(* Logix 5000 project; controller FV vendor 1 type 14 code 217 rev 31.11; software revision 31.00; part 8 of 63 *)
(* tags used below, declared in another part *)
   CWD : CHECKWORD_FLAGS;
   FR_B240 : INT[255];   // DEBOUNCE Debounce Flags
   FR_Delphi_I : DINT[60];
   FR_FILT_PR_PX : PlantItem;   // FILT_PR_PX
   FR_FILT_PR_PX_RawInput : ALIAS FOR RIO_Rack_2:3:I.Data.25;   // FR_FILT_PR_PX
   FR_FILT_TNK_PX : PlantItem;   // FILT_TNK_PX
   FR_FILT_TNK_PX_RawInput : ALIAS FOR RIO_Rack_2:3:I.Data.26;   // FR_FILT_TNK_PX
   FR_FILT_TNLN_PX : PlantItem;   // FILT_TNLN_PX
   FR_FILT_TNLN_PX_RawInput : ALIAS FOR RIO_Rack_2:3:I.Data.27;   // FR_FILT_TNLN_PX
   FR_FRV1_LP01 : PlantItem;   // FRV1_LP01
   FR_FRV1_LP01_RawInput : ALIAS FOR RIO_Rack_2:3:I.Data.13;   // FR_FRV1_LP01
   FR_FV26_HLP01 : PlantItem;   // FV26_HLP01
   FR_FV26_HLP01_RawInput : ALIAS FOR RIO_Rack_2:3:I.Data.0;   // FR_FV26_HLP01
   FR_FV26_LLP01 : PlantItem;   // FV26_LLP01
   FR_FV26_LLP01_RawInput : ALIAS FOR RIO_Rack_2:3:I.Data.1;   // FR_FV26_LLP01
   FR_FV27_HLP01 : PlantItem;   // FV27_HLP01
   FR_FV27_HLP01_RawInput : ALIAS FOR RIO_Rack_2:3:I.Data.2;   // FR_FV27_HLP01
   FR_FV27_LLP01 : PlantItem;   // FV27_LLP01
   FR_FV27_LLP01_RawInput : ALIAS FOR RIO_Rack_2:3:I.Data.3;   // FR_FV27_LLP01
   FR_FV28_HLP01 : PlantItem;   // FV28_HLP01
   FR_FV28_HLP01_RawInput : ALIAS FOR RIO_Rack_2:3:I.Data.4;   // FR_FV28_HLP01
   FR_FV28_LLP01 : PlantItem;   // FV28_LLP01
   FR_FV28_LLP01_RawInput : ALIAS FOR RIO_Rack_2:3:I.Data.5;   // FR_FV28_LLP01
   FR_FV29_HLP01 : PlantItem;   // FV29_HLP01
   FR_FV29_HLP01_RawInput : ALIAS FOR RIO_Rack_2:3:I.Data.6;   // FR_FV29_HLP01
   FR_FV29_LLP01 : PlantItem;   // FV29_LLP01
   FR_FV29_LLP01_RawInput : ALIAS FOR RIO_Rack_2:3:I.Data.7;   // FR_FV29_LLP01
   FR_FV30_HLP01 : PlantItem;   // FV30_HLP01
   FR_FV30_HLP01_RawInput : ALIAS FOR RIO_Rack_2:3:I.Data.8;   // FR_FV30_HLP01
   FR_FV30_LLP01 : PlantItem;   // FV30_LLP01
   FR_FV30_LLP01_RawInput : ALIAS FOR RIO_Rack_2:3:I.Data.9;   // FR_FV30_LLP01
   FR_FV31_HLP01 : PlantItem;   // FV31_HLP01
   FR_FV31_HLP01_RawInput : ALIAS FOR RIO_Rack_2:3:I.Data.10;   // FR_FV31_HLP01
   FR_FV31_LLP01 : PlantItem;   // FV31_LLP01
   FR_FV31_LLP01_RawInput : ALIAS FOR RIO_Rack_2:3:I.Data.11;   // FR_FV31_LLP01
   FR_R3_SW3_3 : PlantItem;   // R3_SW3_3
   FR_R3_SW3_3_RawInput : ALIAS FOR RIO_Rack_2:3:I.Data.14;   // FR_R3_SW3_3 FR_N14[109].2
   FR_T242 : TIMER[255];   // DEBOUNCE
   FR_T243 : TIMER[255];   // DEBOUNCE
   FR_VB4_LP01 : PlantItem;   // VB4_LP01
   FR_VB4_LP01_RawInput : ALIAS FOR RIO_Rack_2:3:I.Data.12;   // FR_VB4_LP01
   FR_YP1_CIPRET : PlantItem;   // YP1_CIPRET
   FR_YP1_CIPRET_RawInput : ALIAS FOR RIO_Rack_2:3:I.Data.24;   // FR_YP1_CIPRET
   FR_YP2_CIPRET : PlantItem;   // YP2_CIPRET
   FR_YP2_CIPRET_RawInput : ALIAS FOR RIO_Rack_2:3:I.Data.22;   // FR_YP2_CIPRET
   FR_YP3_CIPRET : PlantItem;   // YP3_CIPRET
   FR_YP3_CIPRET_RawInput : ALIAS FOR RIO_Rack_2:3:I.Data.23;   // FR_YP3_CIPRET
   One_Second_One_Scan : ALIAS FOR One_Second_1_scan;
(* FR_Common, continued *)

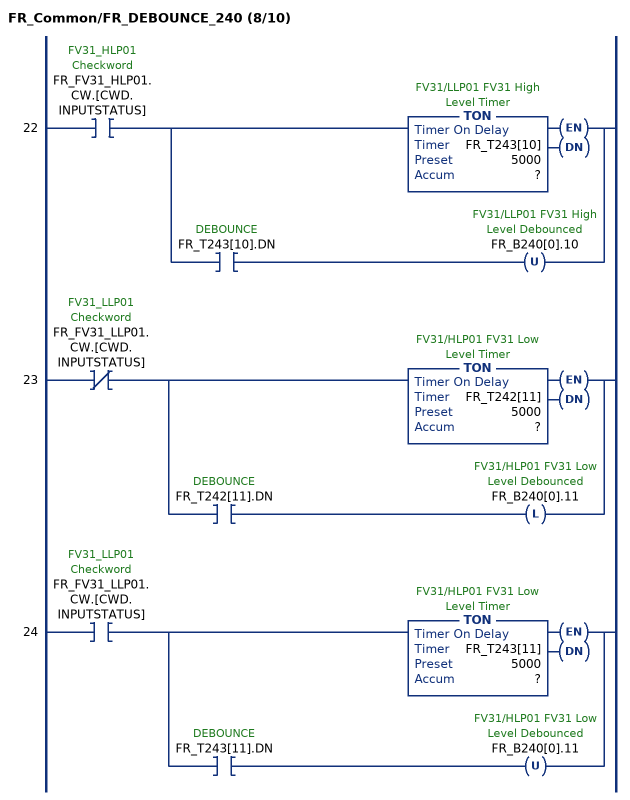
   [picture p70: FR_Common/FR_DEBOUNCE_240 rungs 22-24]
   22: XIC(FR_FV31_HLP01.CW.[CWD.INPUTSTATUS])[TON(FR_T243[10],?,?) ,XIC(FR_T243[10].DN) OTU(FR_B240[0].10) ];
   23: XIO(FR_FV31_LLP01.CW.[CWD.INPUTSTATUS])[TON(FR_T242[11],?,?) ,XIC(FR_T242[11].DN) OTL(FR_B240[0].11) ];
   24: XIC(FR_FV31_LLP01.CW.[CWD.INPUTSTATUS])[TON(FR_T243[11],?,?) ,XIC(FR_T243[11].DN) OTU(FR_B240[0].11) ];
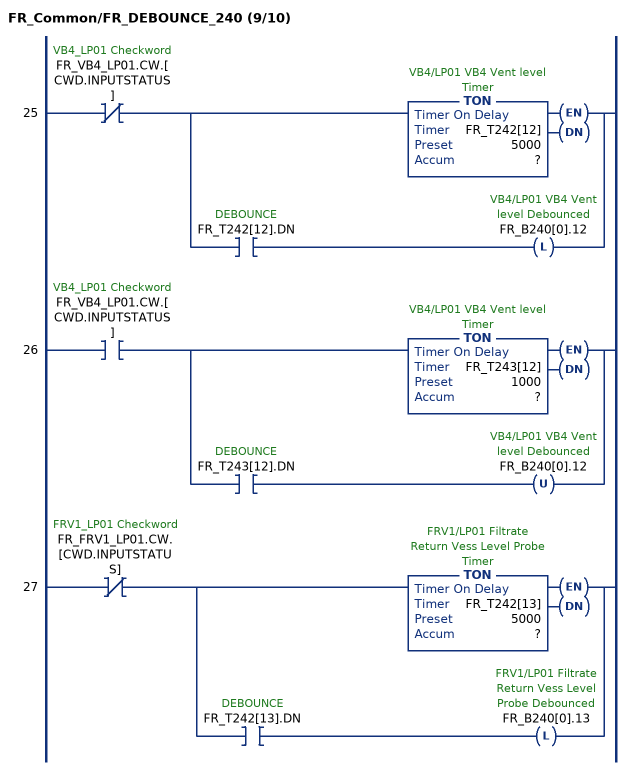
   25: XIO(FR_VB4_LP01.CW.[CWD.INPUTSTATUS])[TON(FR_T242[12],?,?) ,XIC(FR_T242[12].DN) OTL(FR_B240[0].12) ];
   26: XIC(FR_VB4_LP01.CW.[CWD.INPUTSTATUS])[TON(FR_T243[12],?,?) ,XIC(FR_T243[12].DN) OTU(FR_B240[0].12) ];
   27: XIO(FR_FRV1_LP01.CW.[CWD.INPUTSTATUS])[TON(FR_T242[13],?,?) ,XIC(FR_T242[13].DN) OTL(FR_B240[0].13) ];
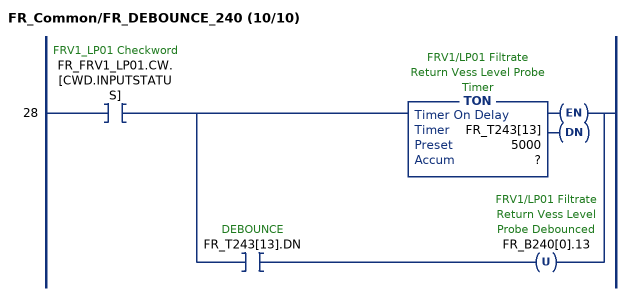
   28: XIC(FR_FRV1_LP01.CW.[CWD.INPUTSTATUS])[TON(FR_T243[13],?,?) ,XIC(FR_T243[13].DN) OTU(FR_B240[0].13) ];
END_ROUTINE

ROUTINE FR_Digital_Inputs   (* ladder *)
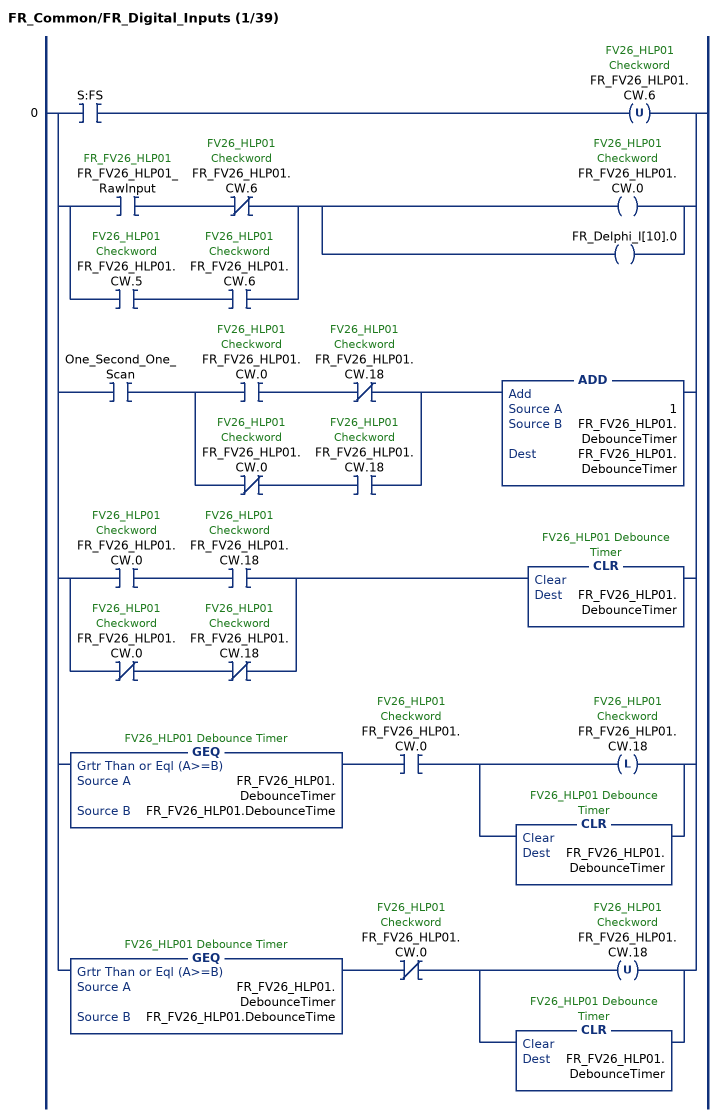
   0: [XIC(S:FS) OTU(FR_FV26_HLP01.CW.6) ,[XIC(FR_FV26_HLP01_RawInput) XIO(FR_FV26_HLP01.CW.6) ,XIC(FR_FV26_HLP01.CW.5) XIC(FR_FV26_HLP01.CW.6) ] [OTE(FR_FV26_HLP01.CW.0) ,OTE(FR_Delphi_I[10].0) ] ,XIC(One_Second_One_Scan) [XIC(FR_FV26_HLP01.CW.0) XIO(FR_FV26_HLP01.CW.18) ,XIO(FR_FV26_HLP01.CW.0) XIC(FR_FV26_HLP01.CW.18) ] ADD(1,FR_FV26_HLP01.DebounceTimer,FR_FV26_HLP01.DebounceTimer) ,[XIC(FR_FV26_HLP01.CW.0) XIC(FR_FV26_HLP01.CW.18) ,XIO(FR_FV26_HLP01.CW.0) XIO(FR_FV26_HLP01.CW.18) ] CLR(FR_FV26_HLP01.DebounceTimer) ,GEQ(FR_FV26_HLP01.DebounceTimer,FR_FV26_HLP01.DebounceTime) XIC(FR_FV26_HLP01.CW.0) [OTL(FR_FV26_HLP01.CW.18) ,CLR(FR_FV26_HLP01.DebounceTimer) ] ,GEQ(FR_FV26_HLP01.DebounceTimer,FR_FV26_HLP01.DebounceTime) XIO(FR_FV26_HLP01.CW.0) [OTU(FR_FV26_HLP01.CW.18) ,CLR(FR_FV26_HLP01.DebounceTimer) ] ];
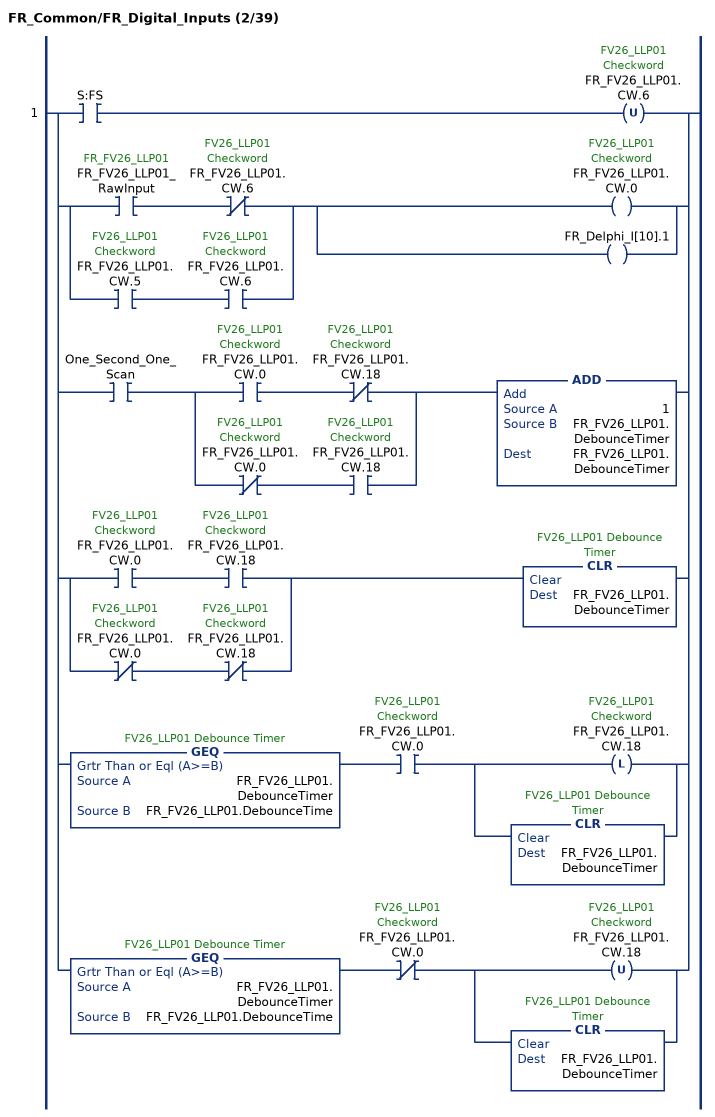
   1: [XIC(S:FS) OTU(FR_FV26_LLP01.CW.6) ,[XIC(FR_FV26_LLP01_RawInput) XIO(FR_FV26_LLP01.CW.6) ,XIC(FR_FV26_LLP01.CW.5) XIC(FR_FV26_LLP01.CW.6) ] [OTE(FR_FV26_LLP01.CW.0) ,OTE(FR_Delphi_I[10].1) ] ,XIC(One_Second_One_Scan) [XIC(FR_FV26_LLP01.CW.0) XIO(FR_FV26_LLP01.CW.18) ,XIO(FR_FV26_LLP01.CW.0) XIC(FR_FV26_LLP01.CW.18) ] ADD(1,FR_FV26_LLP01.DebounceTimer,FR_FV26_LLP01.DebounceTimer) ,[XIC(FR_FV26_LLP01.CW.0) XIC(FR_FV26_LLP01.CW.18) ,XIO(FR_FV26_LLP01.CW.0) XIO(FR_FV26_LLP01.CW.18) ] CLR(FR_FV26_LLP01.DebounceTimer) ,GEQ(FR_FV26_LLP01.DebounceTimer,FR_FV26_LLP01.DebounceTime) XIC(FR_FV26_LLP01.CW.0) [OTL(FR_FV26_LLP01.CW.18) ,CLR(FR_FV26_LLP01.DebounceTimer) ] ,GEQ(FR_FV26_LLP01.DebounceTimer,FR_FV26_LLP01.DebounceTime) XIO(FR_FV26_LLP01.CW.0) [OTU(FR_FV26_LLP01.CW.18) ,CLR(FR_FV26_LLP01.DebounceTimer) ] ];
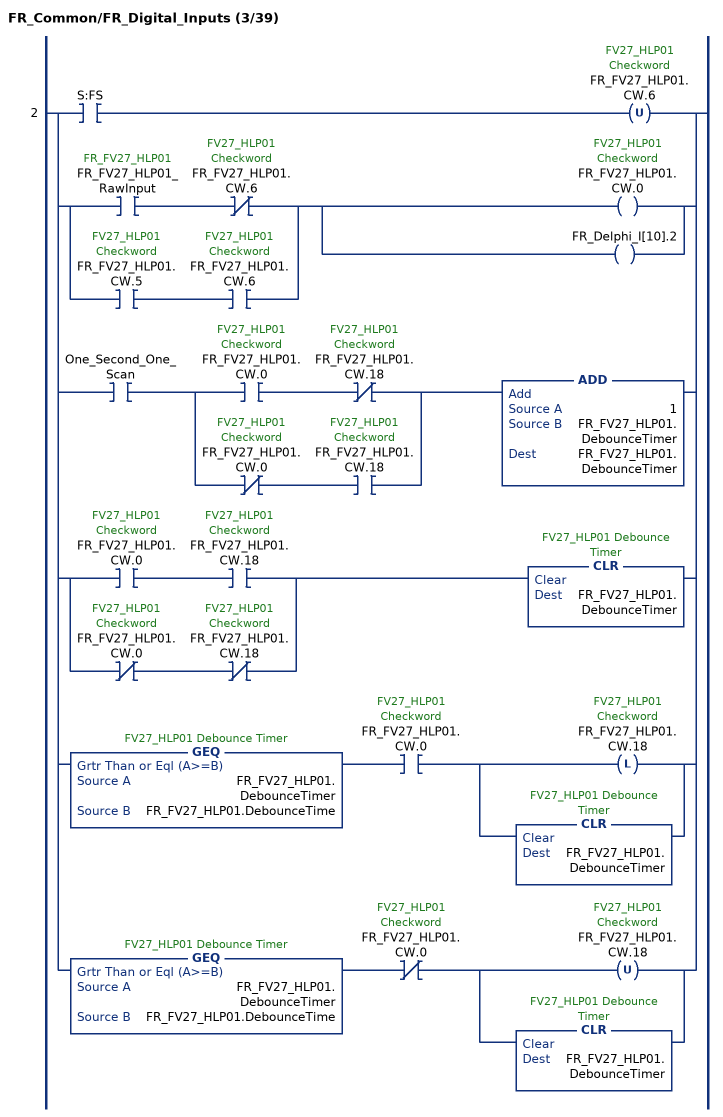
   2: [XIC(S:FS) OTU(FR_FV27_HLP01.CW.6) ,[XIC(FR_FV27_HLP01_RawInput) XIO(FR_FV27_HLP01.CW.6) ,XIC(FR_FV27_HLP01.CW.5) XIC(FR_FV27_HLP01.CW.6) ] [OTE(FR_FV27_HLP01.CW.0) ,OTE(FR_Delphi_I[10].2) ] ,XIC(One_Second_One_Scan) [XIC(FR_FV27_HLP01.CW.0) XIO(FR_FV27_HLP01.CW.18) ,XIO(FR_FV27_HLP01.CW.0) XIC(FR_FV27_HLP01.CW.18) ] ADD(1,FR_FV27_HLP01.DebounceTimer,FR_FV27_HLP01.DebounceTimer) ,[XIC(FR_FV27_HLP01.CW.0) XIC(FR_FV27_HLP01.CW.18) ,XIO(FR_FV27_HLP01.CW.0) XIO(FR_FV27_HLP01.CW.18) ] CLR(FR_FV27_HLP01.DebounceTimer) ,GEQ(FR_FV27_HLP01.DebounceTimer,FR_FV27_HLP01.DebounceTime) XIC(FR_FV27_HLP01.CW.0) [OTL(FR_FV27_HLP01.CW.18) ,CLR(FR_FV27_HLP01.DebounceTimer) ] ,GEQ(FR_FV27_HLP01.DebounceTimer,FR_FV27_HLP01.DebounceTime) XIO(FR_FV27_HLP01.CW.0) [OTU(FR_FV27_HLP01.CW.18) ,CLR(FR_FV27_HLP01.DebounceTimer) ] ];
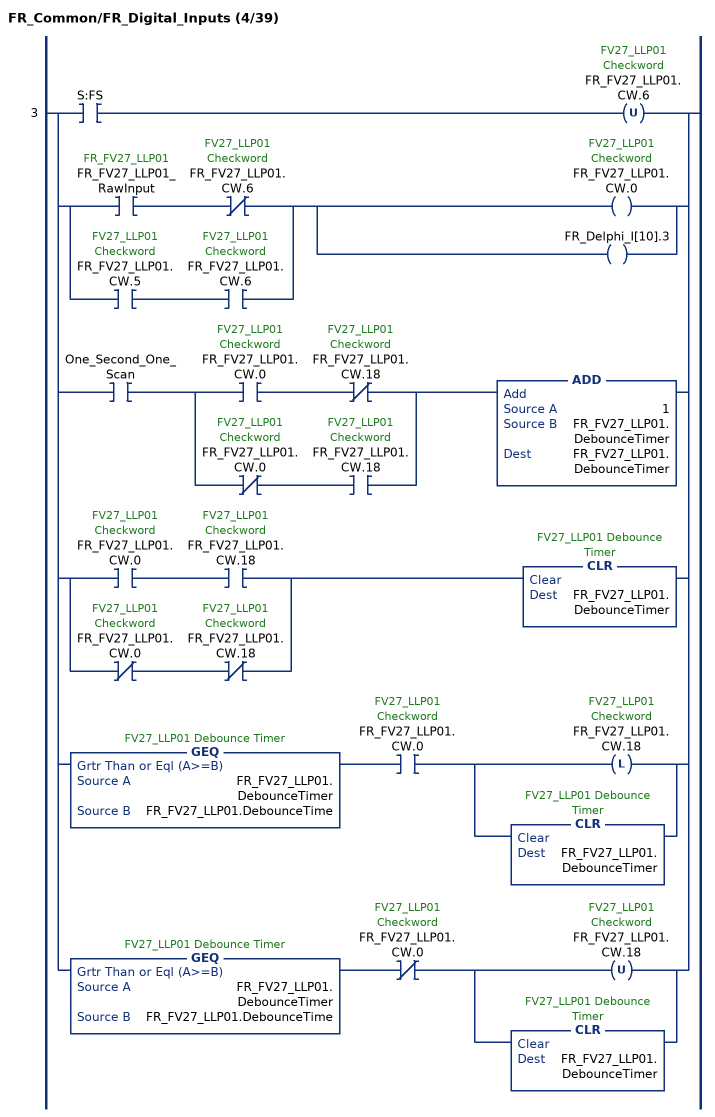
   3: [XIC(S:FS) OTU(FR_FV27_LLP01.CW.6) ,[XIC(FR_FV27_LLP01_RawInput) XIO(FR_FV27_LLP01.CW.6) ,XIC(FR_FV27_LLP01.CW.5) XIC(FR_FV27_LLP01.CW.6) ] [OTE(FR_FV27_LLP01.CW.0) ,OTE(FR_Delphi_I[10].3) ] ,XIC(One_Second_One_Scan) [XIC(FR_FV27_LLP01.CW.0) XIO(FR_FV27_LLP01.CW.18) ,XIO(FR_FV27_LLP01.CW.0) XIC(FR_FV27_LLP01.CW.18) ] ADD(1,FR_FV27_LLP01.DebounceTimer,FR_FV27_LLP01.DebounceTimer) ,[XIC(FR_FV27_LLP01.CW.0) XIC(FR_FV27_LLP01.CW.18) ,XIO(FR_FV27_LLP01.CW.0) XIO(FR_FV27_LLP01.CW.18) ] CLR(FR_FV27_LLP01.DebounceTimer) ,GEQ(FR_FV27_LLP01.DebounceTimer,FR_FV27_LLP01.DebounceTime) XIC(FR_FV27_LLP01.CW.0) [OTL(FR_FV27_LLP01.CW.18) ,CLR(FR_FV27_LLP01.DebounceTimer) ] ,GEQ(FR_FV27_LLP01.DebounceTimer,FR_FV27_LLP01.DebounceTime) XIO(FR_FV27_LLP01.CW.0) [OTU(FR_FV27_LLP01.CW.18) ,CLR(FR_FV27_LLP01.DebounceTimer) ] ];
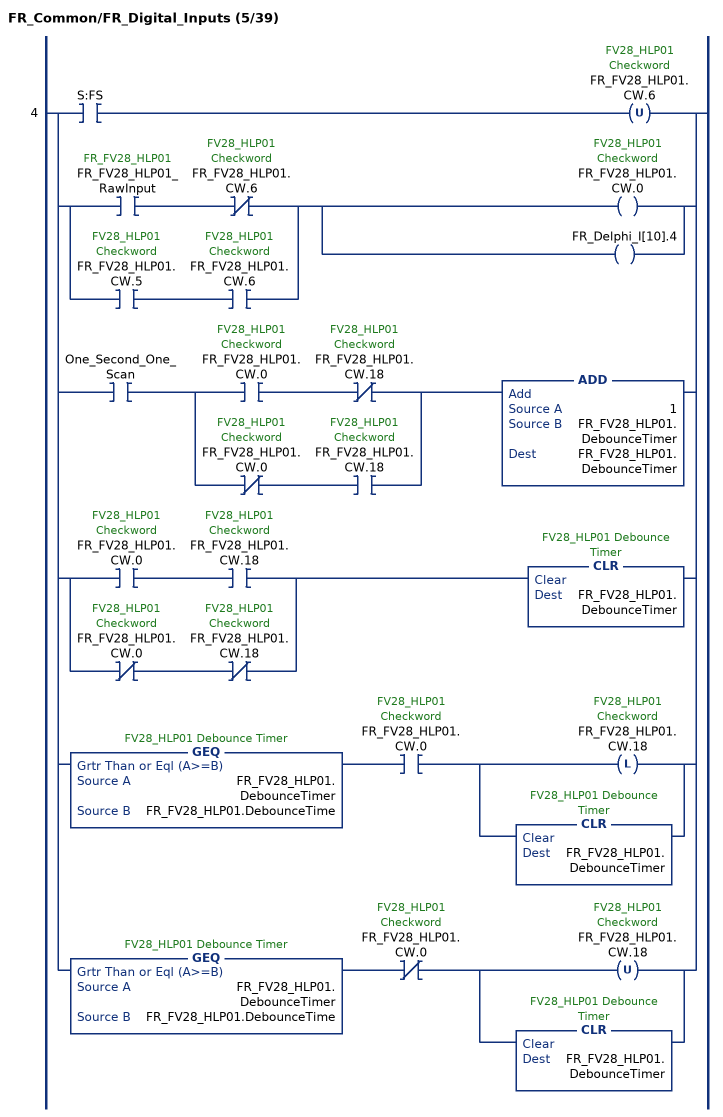
   4: [XIC(S:FS) OTU(FR_FV28_HLP01.CW.6) ,[XIC(FR_FV28_HLP01_RawInput) XIO(FR_FV28_HLP01.CW.6) ,XIC(FR_FV28_HLP01.CW.5) XIC(FR_FV28_HLP01.CW.6) ] [OTE(FR_FV28_HLP01.CW.0) ,OTE(FR_Delphi_I[10].4) ] ,XIC(One_Second_One_Scan) [XIC(FR_FV28_HLP01.CW.0) XIO(FR_FV28_HLP01.CW.18) ,XIO(FR_FV28_HLP01.CW.0) XIC(FR_FV28_HLP01.CW.18) ] ADD(1,FR_FV28_HLP01.DebounceTimer,FR_FV28_HLP01.DebounceTimer) ,[XIC(FR_FV28_HLP01.CW.0) XIC(FR_FV28_HLP01.CW.18) ,XIO(FR_FV28_HLP01.CW.0) XIO(FR_FV28_HLP01.CW.18) ] CLR(FR_FV28_HLP01.DebounceTimer) ,GEQ(FR_FV28_HLP01.DebounceTimer,FR_FV28_HLP01.DebounceTime) XIC(FR_FV28_HLP01.CW.0) [OTL(FR_FV28_HLP01.CW.18) ,CLR(FR_FV28_HLP01.DebounceTimer) ] ,GEQ(FR_FV28_HLP01.DebounceTimer,FR_FV28_HLP01.DebounceTime) XIO(FR_FV28_HLP01.CW.0) [OTU(FR_FV28_HLP01.CW.18) ,CLR(FR_FV28_HLP01.DebounceTimer) ] ];
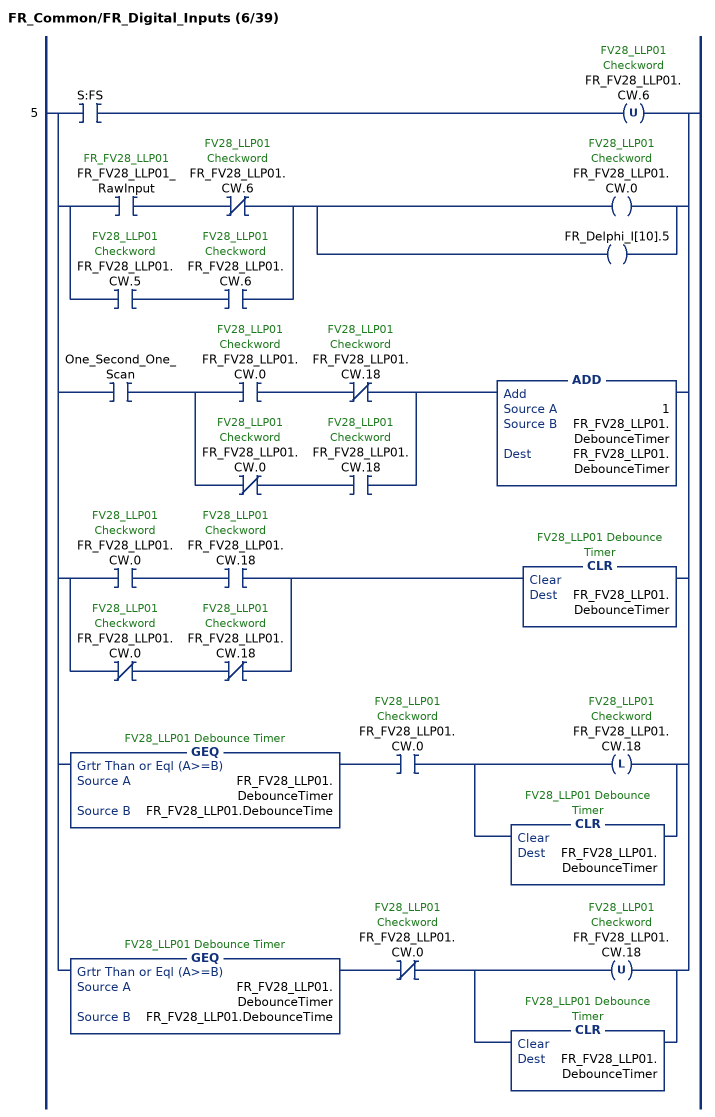
   5: [XIC(S:FS) OTU(FR_FV28_LLP01.CW.6) ,[XIC(FR_FV28_LLP01_RawInput) XIO(FR_FV28_LLP01.CW.6) ,XIC(FR_FV28_LLP01.CW.5) XIC(FR_FV28_LLP01.CW.6) ] [OTE(FR_FV28_LLP01.CW.0) ,OTE(FR_Delphi_I[10].5) ] ,XIC(One_Second_One_Scan) [XIC(FR_FV28_LLP01.CW.0) XIO(FR_FV28_LLP01.CW.18) ,XIO(FR_FV28_LLP01.CW.0) XIC(FR_FV28_LLP01.CW.18) ] ADD(1,FR_FV28_LLP01.DebounceTimer,FR_FV28_LLP01.DebounceTimer) ,[XIC(FR_FV28_LLP01.CW.0) XIC(FR_FV28_LLP01.CW.18) ,XIO(FR_FV28_LLP01.CW.0) XIO(FR_FV28_LLP01.CW.18) ] CLR(FR_FV28_LLP01.DebounceTimer) ,GEQ(FR_FV28_LLP01.DebounceTimer,FR_FV28_LLP01.DebounceTime) XIC(FR_FV28_LLP01.CW.0) [OTL(FR_FV28_LLP01.CW.18) ,CLR(FR_FV28_LLP01.DebounceTimer) ] ,GEQ(FR_FV28_LLP01.DebounceTimer,FR_FV28_LLP01.DebounceTime) XIO(FR_FV28_LLP01.CW.0) [OTU(FR_FV28_LLP01.CW.18) ,CLR(FR_FV28_LLP01.DebounceTimer) ] ];
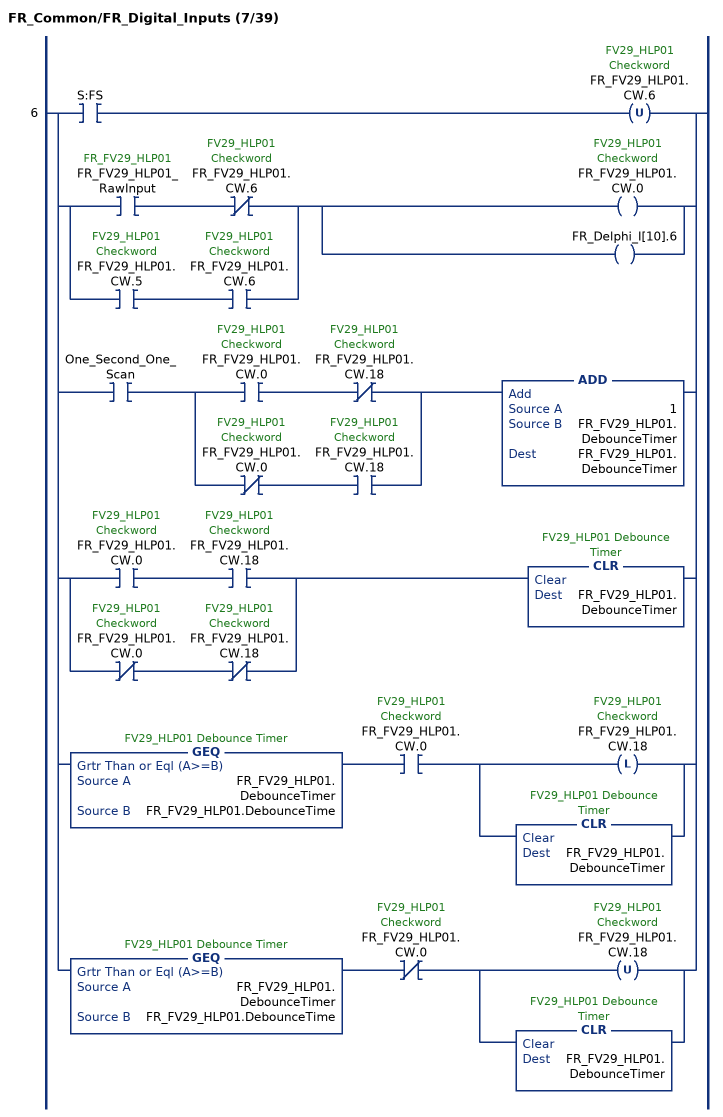
   6: [XIC(S:FS) OTU(FR_FV29_HLP01.CW.6) ,[XIC(FR_FV29_HLP01_RawInput) XIO(FR_FV29_HLP01.CW.6) ,XIC(FR_FV29_HLP01.CW.5) XIC(FR_FV29_HLP01.CW.6) ] [OTE(FR_FV29_HLP01.CW.0) ,OTE(FR_Delphi_I[10].6) ] ,XIC(One_Second_One_Scan) [XIC(FR_FV29_HLP01.CW.0) XIO(FR_FV29_HLP01.CW.18) ,XIO(FR_FV29_HLP01.CW.0) XIC(FR_FV29_HLP01.CW.18) ] ADD(1,FR_FV29_HLP01.DebounceTimer,FR_FV29_HLP01.DebounceTimer) ,[XIC(FR_FV29_HLP01.CW.0) XIC(FR_FV29_HLP01.CW.18) ,XIO(FR_FV29_HLP01.CW.0) XIO(FR_FV29_HLP01.CW.18) ] CLR(FR_FV29_HLP01.DebounceTimer) ,GEQ(FR_FV29_HLP01.DebounceTimer,FR_FV29_HLP01.DebounceTime) XIC(FR_FV29_HLP01.CW.0) [OTL(FR_FV29_HLP01.CW.18) ,CLR(FR_FV29_HLP01.DebounceTimer) ] ,GEQ(FR_FV29_HLP01.DebounceTimer,FR_FV29_HLP01.DebounceTime) XIO(FR_FV29_HLP01.CW.0) [OTU(FR_FV29_HLP01.CW.18) ,CLR(FR_FV29_HLP01.DebounceTimer) ] ];
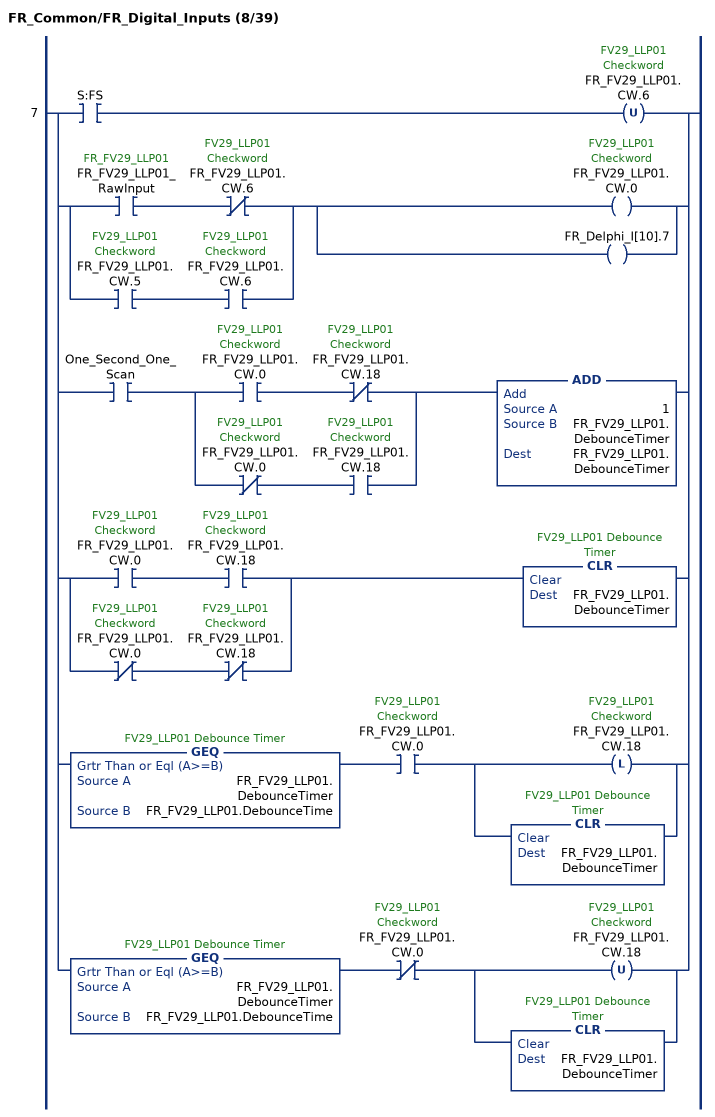
   7: [XIC(S:FS) OTU(FR_FV29_LLP01.CW.6) ,[XIC(FR_FV29_LLP01_RawInput) XIO(FR_FV29_LLP01.CW.6) ,XIC(FR_FV29_LLP01.CW.5) XIC(FR_FV29_LLP01.CW.6) ] [OTE(FR_FV29_LLP01.CW.0) ,OTE(FR_Delphi_I[10].7) ] ,XIC(One_Second_One_Scan) [XIC(FR_FV29_LLP01.CW.0) XIO(FR_FV29_LLP01.CW.18) ,XIO(FR_FV29_LLP01.CW.0) XIC(FR_FV29_LLP01.CW.18) ] ADD(1,FR_FV29_LLP01.DebounceTimer,FR_FV29_LLP01.DebounceTimer) ,[XIC(FR_FV29_LLP01.CW.0) XIC(FR_FV29_LLP01.CW.18) ,XIO(FR_FV29_LLP01.CW.0) XIO(FR_FV29_LLP01.CW.18) ] CLR(FR_FV29_LLP01.DebounceTimer) ,GEQ(FR_FV29_LLP01.DebounceTimer,FR_FV29_LLP01.DebounceTime) XIC(FR_FV29_LLP01.CW.0) [OTL(FR_FV29_LLP01.CW.18) ,CLR(FR_FV29_LLP01.DebounceTimer) ] ,GEQ(FR_FV29_LLP01.DebounceTimer,FR_FV29_LLP01.DebounceTime) XIO(FR_FV29_LLP01.CW.0) [OTU(FR_FV29_LLP01.CW.18) ,CLR(FR_FV29_LLP01.DebounceTimer) ] ];
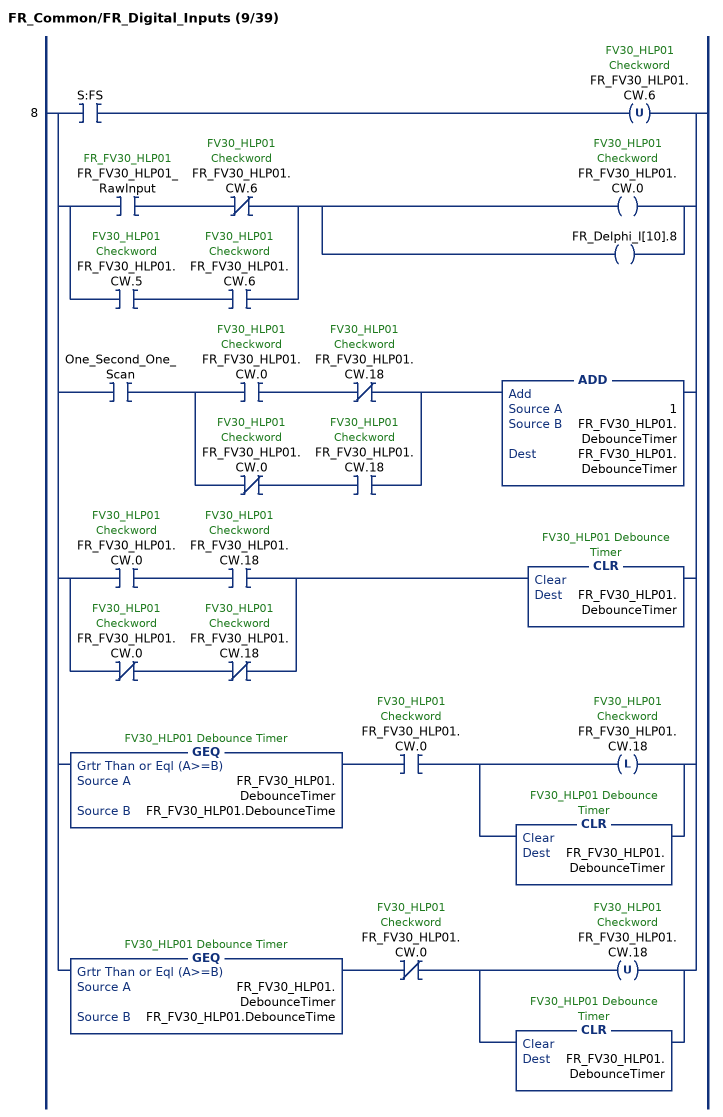
   8: [XIC(S:FS) OTU(FR_FV30_HLP01.CW.6) ,[XIC(FR_FV30_HLP01_RawInput) XIO(FR_FV30_HLP01.CW.6) ,XIC(FR_FV30_HLP01.CW.5) XIC(FR_FV30_HLP01.CW.6) ] [OTE(FR_FV30_HLP01.CW.0) ,OTE(FR_Delphi_I[10].8) ] ,XIC(One_Second_One_Scan) [XIC(FR_FV30_HLP01.CW.0) XIO(FR_FV30_HLP01.CW.18) ,XIO(FR_FV30_HLP01.CW.0) XIC(FR_FV30_HLP01.CW.18) ] ADD(1,FR_FV30_HLP01.DebounceTimer,FR_FV30_HLP01.DebounceTimer) ,[XIC(FR_FV30_HLP01.CW.0) XIC(FR_FV30_HLP01.CW.18) ,XIO(FR_FV30_HLP01.CW.0) XIO(FR_FV30_HLP01.CW.18) ] CLR(FR_FV30_HLP01.DebounceTimer) ,GEQ(FR_FV30_HLP01.DebounceTimer,FR_FV30_HLP01.DebounceTime) XIC(FR_FV30_HLP01.CW.0) [OTL(FR_FV30_HLP01.CW.18) ,CLR(FR_FV30_HLP01.DebounceTimer) ] ,GEQ(FR_FV30_HLP01.DebounceTimer,FR_FV30_HLP01.DebounceTime) XIO(FR_FV30_HLP01.CW.0) [OTU(FR_FV30_HLP01.CW.18) ,CLR(FR_FV30_HLP01.DebounceTimer) ] ];